   Warranty conditions, liability, AND support -
      IF the application has been made available free OF charge, the following applies:
      * We DO NOT provide a warranty FOR Any OF the information contained in this document.
      * All other rights AND claims against Siemens AG irrespective OF legal basis are excluded. In particular claims FOR damages against Siemens AG 
      in the CASE OF Product outage, downtime, loss OF profit, either directly, indirectly OR consequential damage are excluded.
      * This does NOT apply when liability is compulsory BY law, e. g. in the CASE OF the Product liability act, premeditation, an act OF gross negligence 
      BY superiors AND managerial staff OF Siemens AG OR in cases OF fraudulent concealment OF defects.
      * This limitation OF liability also applies TO sub-contractors, suppliers, delegates, superiors AND managerial staff OF Siemens AG.
      German law shall apply TO this agreement FOR customers with head offices in Germany; Swiss law FOR customers with head offices outside Germany. 
      Application OF the United Nations Convention on Contracts FOR the International Sale OF Goods as OF 11.04.1980 (CISG) is excluded.
   *)

   // ===========================================================================
   //  Begin the LOGIC section:
   //  

    #temp_UDint := 0;

   IF IS_ARRAY(#Array_ToBe_Sized) THEN                             // Is this a valid array?
       #temp_UDint := CountOfElements(#Array_ToBe_Sized);          // Determine the length of the array...
   END_IF;

   #ArraySize := UDINT_TO_INT(#temp_UDint);

   // End of Main Logic Section 
   ENO := true;   // Set the ENO output
END_FUNCTION

(* ===== HMI "HMI_RT_1" =====
system functions are stored by id; their names below are inferred from use

HMI tags "Default tag table"
   "bo_PreviousPage_pressed" : Bool, internal
   "bo_NextPage_pressed" : Bool, internal

ScreenModuleEditorView "typ_ThirdLevelNavigation" 165x50
   Button "Btn_NextPage" at 115,0 size 50x50; TextOff 'Text'; PictureOff "Right_transparent_48x48"
      on Press: function_b14e0dd5("bo_NextPage_pressed", 0)
      Appearance <- "bo_NextPage_pressed"
   Button "btn_PreviousPage" at 0,0 size 50x50; TextOff 'Text'; PictureOff "Left_transparent_48x48"
      on Press: function_b14e0dd5("bo_PreviousPage_pressed", 0)
      Appearance <- "bo_PreviousPage_pressed"
   TextField "txt_actualID" at 55,11 size 28x27; Text '11'
   TextField "txt_maximum _ID" at 82,11 size 28x27; Text '11'
   TextField "txt_Backslash" at 76,11 size 14x27; Text '/'
   GraphicView "pic_transparent_previous" at 0,0 size 50x50; Picture "btn-disabled-50x50"
      Visibility <- "bo_PreviousActive"
   GraphicView "pic_transparent_next" at 115,0 size 50x50; Picture "btn-disabled-50x50"
      Visibility <- "bo_NextActive"
*)

(* ===== HMI "HMI_RT_1" =====

ScreenModuleEditorView "fcpOmacTime" 490x26
   IOField "valOutputModeName" at 0,0 size 151x26; FormatPattern ??????????????????
      ProcessValue <- "ModeName"
   IOField "valOutputCurrentTime" at 150,0 size 101x26; FormatPattern 999999999
      ProcessValue <- "CurrentTime"
   IOField "ValOutputCumulativeTime" at 250,0 size 101x26; FormatPattern 999999999
      ProcessValue <- "CumulativeTime"
   Bar "valOutputCumuliativeTimePercent" at 355,5 size 131x16; MinimumValue 0; MaximumValue 100
      ProcessValue <- "CumulativeTime"
      MaximumValue <- "TimeOverAll"
*)

(* ===== HMI "HMI_RT_1" =====
system functions are stored by id; their names below are inferred from use

HMI tags "Standard-Variablentabelle"
   "bo_Topic01BtnPressed" : Bool, internal
   "bo_Topic02BtnPressed" : Bool, internal
   "bo_Topic03BtnPressed" : Bool, internal
   "bo_Topic04BtnPressed" : Bool, internal
   "bo_Topic05BtnPressed" : Bool, internal
   "bo_Topic06BtnPressed" : Bool, internal
   "bo_Topic07BtnPressed" : Bool, internal
   "bo_Topic08BtnPressed" : Bool, internal
   "bo_Topic09BtnPressed" : Bool, internal
   "bo_Topic10BtnPressed" : Bool, internal
   "bo_Topic11BtnPressed" : Bool, internal
   "bo_Topic12BtnPressed" : Bool, internal
   "bo_Topic13BtnPressed" : Bool, internal
   "bo_Topic14BtnPressed" : Bool, internal
   "bo_Topic15BtnPressed" : Bool, internal
   "bo_Topic16BtnPressed" : Bool, internal
   "bo_Topic17BtnPressed" : Bool, internal
   "bo_Topic18BtnPressed" : Bool, internal
   "bo_Topic19BtnPressed" : Bool, internal
   "bo_Topic20BtnPressed" : Bool, internal
   "bo_Topic21BtnPressed" : Bool, internal
   "bo_Topic22BtnPressed" : Bool, internal
   "bo_Topic23BtnPressed" : Bool, internal
   "bo_Topic24BtnPressed" : Bool, internal
   "i16_configReg" : Int, internal   // Combination of actual showed LvL and input configuration of used Register; To show active Register
   "i16_LvL_Shown" : Int, internal   // number of actual showed LvL
   "i16_SaveScreenNo" : Int, internal   // Save actual Screen Number
   "i16_RegShown" : Int, internal   // Combination of actual active Register and actual active LvL; to show the active Register
   "bo_NextTopicLvL1" : Int, internal
   "i16_InputScreenID" : Int, internal   // help Variable
   "i16_Input_maxReg" : Int, internal   // help Variable
   "i16_RegNo" : Int, internal   // Active Register number;Value 1-24
   "bo_PreviousPageBtnPressed" : Bool, internal

ScreenModuleEditorView "fcpSecondLevelNavigation" 1270x615
   Rectangle "rec_Topic_001.0" at 207,42 size 1063x62
      Visibility <- "i16_RegShown"
   Rectangle "rec_Topic_002.0" at 207,109 size 1063x62
      Visibility <- "i16_RegShown"
   Rectangle "rec_Topic_003.0" at 207,176 size 1063x62
      Visibility <- "i16_RegShown"
   Rectangle "rec_Topic_004.0" at 207,243 size 1063x62
      Visibility <- "i16_RegShown"
   Rectangle "rec_Topic_005.0" at 207,310 size 1063x62
      Visibility <- "i16_RegShown"
   Rectangle "rec_Topic_006.0" at 207,377 size 1063x62
      Visibility <- "i16_RegShown"
   Rectangle "rec_Topic_007.0" at 207,444 size 1063x62
      Visibility <- "i16_RegShown"
   Rectangle "rec_Topic_008.0" at 207,511 size 1063x62
      Visibility <- "i16_RegShown"
   TextField "txt_Topic_001.0_Textfield" at 1100,42 size 170x62; Text 'Thema 001.0 / Topic 001.0'
      Visibility <- "i16_configReg"
      Appearance <- "i16_RegShown"
   Button "btn_Topic_001.0_Button" at 1100,42 size 170x62; TextOff 'Text'
      on Release: "sub_TabLvL"()
      on Press: function_b14e0dd5("bo_Topic01BtnPressed", 0)
      Visibility <- "i16_configReg"
   TextField "txt_Topic_002.0_Textfield" at 1100,109 size 170x62; Text 'Thema 002.0 / Topic 002.0'
      Visibility <- "i16_configReg"
      Appearance <- "i16_RegShown"
   Button "btn_Topic_002.0_Button" at 1100,109 size 170x62; TextOff 'Text'
      on Release: "sub_TabLvL"()
      on Press: function_b14e0dd5("bo_Topic02BtnPressed", 0)
      Visibility <- "i16_configReg"
   TextField "txt_Topic_003.0_Textfield" at 1100,176 size 170x62; Text 'Thema 003.0 / Topic 003.0'
      Visibility <- "i16_configReg"
      Appearance <- "i16_RegShown"
   Button "btn_Topic_003.0_Button" at 1100,176 size 170x62; TextOff 'Text'
      on Release: "sub_TabLvL"()
      on Press: function_b14e0dd5("bo_Topic03BtnPressed", 0)
      Visibility <- "i16_configReg"
   TextField "txt_Topic_004.0_Textfield" at 1100,243 size 170x62; Text 'Thema 004.0 / Topic 004.0'
      Visibility <- "i16_configReg"
      Appearance <- "i16_RegShown"
   Button "btn_Topic_004.0_Button" at 1100,243 size 170x62; TextOff 'Text'
      on Release: "sub_TabLvL"()
      on Press: function_b14e0dd5("bo_Topic04BtnPressed", 0)
      Visibility <- "i16_configReg"
   TextField "txt_Topic_005.0_Textfield" at 1100,310 size 170x62; Text 'Thema 005.0 / Topic 005.0'
      Visibility <- "i16_configReg"
      Appearance <- "i16_RegShown"
   Button "btn_Topic_005.0_Button" at 1100,310 size 170x62; TextOff 'Text'
      on Release: "sub_TabLvL"()
      on Press: function_b14e0dd5("bo_Topic05BtnPressed", 0)
      Visibility <- "i16_configReg"
   TextField "txt_Topic_006.0_Textfield" at 1100,377 size 170x62; Text 'Thema 006.0 / Topic 006.0 / Topic 005.0'
      Visibility <- "i16_configReg"
      Appearance <- "i16_RegShown"
   Button "btn_Topic_006.0_Button" at 1100,377 size 170x62; TextOff 'Text'
      on Release: "sub_TabLvL"()
      on Press: function_b14e0dd5("bo_Topic06BtnPressed", 0)
      Visibility <- "i16_configReg"
   TextField "txt_Topic_007.0_Textfield" at 1100,444 size 170x62; Text 'Thema 007.0 / Topic 007.0 / Topic 005.0'
      Visibility <- "i16_configReg"
      Appearance <- "i16_RegShown"
   Button "btn_Topic_007.0_Button" at 1100,444 size 170x62; TextOff 'Text'
      on Release: "sub_TabLvL"()
      on Press: function_b14e0dd5("bo_Topic07BtnPressed", 0)
      Visibility <- "i16_configReg"
   TextField "txt_Topic_008.0_Textfield" at 1100,511 size 170x62; Text 'Thema 007.0 / Topic 008.0 / Topic 005.0'
      Visibility <- "i16_configReg"
      Appearance <- "i16_RegShown"
   Button "btn_Topic_008.0_Button" at 1100,511 size 170x62; TextOff 'Text'
      on Release: "sub_TabLvL"()
      on Press: function_b14e0dd5("bo_Topic08BtnPressed", 0)
      Visibility <- "i16_configReg"
   Rectangle "rec_Topic_001.0_RectangleLight" at 1100,42 size 170x62
      Visibility <- "i16_configReg"
      Appearance <- "bo_Topic01BtnPressed"
   Rectangle "rec_Topic_002.0_RectangleLight" at 1100,109 size 170x62
      Visibility <- "i16_configReg"
      Appearance <- "bo_Topic02BtnPressed"
   Rectangle "rec_Topic_003.0_RectangleLight" at 1100,176 size 170x62
      Visibility <- "i16_configReg"
      Appearance <- "bo_Topic03BtnPressed"
   Rectangle "rec_Topic_004.0_RectangleLight" at 1100,243 size 170x62
      Visibility <- "i16_configReg"
      Appearance <- "bo_Topic04BtnPressed"
   Rectangle "rec_Topic_005.0_RectangleLight" at 1100,310 size 170x62
      Visibility <- "i16_configReg"
      Appearance <- "bo_Topic05BtnPressed"
   Rectangle "rec_Topic_006.0_RectangleLight" at 1100,377 size 170x62
      Visibility <- "i16_configReg"
      Appearance <- "bo_Topic06BtnPressed"
   Rectangle "rec_Topic_007.0_RectangleLight" at 1100,444 size 170x62
      Visibility <- "i16_configReg"
      Appearance <- "bo_Topic07BtnPressed"
   Rectangle "rec_Topic_008.0_RectangleLight" at 1100,511 size 170x62
      Visibility <- "i16_configReg"
      Appearance <- "bo_Topic08BtnPressed"
   Rectangle "rec_Topic_009.0_RectangleLight" at 1100,42 size 170x62
      Visibility <- "i16_configReg"
      Appearance <- "bo_Topic09BtnPressed"
   Rectangle "rec_Topic_010.0_RectangleLight" at 1100,109 size 170x62
      Visibility <- "i16_configReg"
      Appearance <- "bo_Topic10BtnPressed"
   Rectangle "rec_Topic_011.0_RectangleLight" at 1100,176 size 170x62
      Visibility <- "i16_configReg"
      Appearance <- "bo_Topic11BtnPressed"
   Rectangle "rec_Topic_012.0_RectangleLight" at 1100,243 size 170x62
      Visibility <- "i16_configReg"
      Appearance <- "bo_Topic12BtnPressed"
   Rectangle "rec_Topic_013.0_RectangleLight" at 1100,310 size 170x62
      Visibility <- "i16_configReg"
      Appearance <- "bo_Topic13BtnPressed"
   Rectangle "rec_Topic_014.0_RectangleLight" at 1100,377 size 170x62
      Visibility <- "i16_configReg"
      Appearance <- "bo_Topic14BtnPressed"
   Rectangle "rec_Topic_015.0_RectangleLight" at 1100,444 size 170x62
      Visibility <- "i16_configReg"
      Appearance <- "bo_Topic15BtnPressed"
   Rectangle "rec_Topic_016.0_RectangleLight" at 1100,511 size 170x62
      Visibility <- "i16_configReg"
      Appearance <- "bo_Topic16BtnPressed"
   Rectangle "rec_Topic_009.0" at 207,42 size 1063x62
      Visibility <- "i16_RegShown"
   Rectangle "rec_Topic_010.0" at 207,109 size 1063x62
      Visibility <- "i16_RegShown"
   Rectangle "rec_Topic_011.0" at 207,176 size 1063x62
      Visibility <- "i16_RegShown"
   Rectangle "rec_Topic_012.0" at 207,243 size 1063x62
      Visibility <- "i16_RegShown"
   Rectangle "rec_Topic_013.0" at 207,310 size 1063x62
      Visibility <- "i16_RegShown"
   Rectangle "rec_Topic_014.0" at 207,377 size 1063x62
      Visibility <- "i16_RegShown"
   Rectangle "rec_Topic_015.0" at 207,444 size 1063x62
      Visibility <- "i16_RegShown"
   Rectangle "rec_Topic_016.0" at 207,511 size 1063x62
      Visibility <- "i16_RegShown"
   Rectangle "rec_Topic_017.0_RectangleLight" at 1100,42 size 170x62
      Visibility <- "i16_configReg"
      Appearance <- "bo_Topic17BtnPressed"
   Rectangle "rec_Topic_018.0_RectangleLight" at 1100,109 size 170x62
      Visibility <- "i16_configReg"
      Appearance <- "bo_Topic18BtnPressed"
   Rectangle "rec_Topic_019.0_RectangleLight" at 1100,176 size 170x62
      Visibility <- "i16_configReg"
      Appearance <- "bo_Topic19BtnPressed"
   Rectangle "rec_Topic_020.0_RectangleLight" at 1100,243 size 170x62
      Visibility <- "i16_configReg"
      Appearance <- "bo_Topic20BtnPressed"
   Rectangle "rec_Topic_021.0_RectangleLight" at 1100,310 size 170x62
      Visibility <- "i16_configReg"
      Appearance <- "bo_Topic21BtnPressed"
   Rectangle "rec_Topic_022.0_RectangleLight" at 1100,377 size 170x62
      Visibility <- "i16_configReg"
      Appearance <- "bo_Topic22BtnPressed"
   Rectangle "rec_Topic_023.0_RectangleLight" at 1100,444 size 170x62
      Visibility <- "i16_configReg"
      Appearance <- "bo_Topic23BtnPressed"
   Rectangle "rec_Topic_024.0_RectangleLight" at 1100,511 size 170x62
      Visibility <- "i16_configReg"
      Appearance <- "bo_Topic24BtnPressed"
   Rectangle "rec_Topic_017.0" at 207,42 size 1063x62
      Visibility <- "i16_RegShown"
   Rectangle "rec_Topic_018.0" at 207,109 size 1063x62
      Visibility <- "i16_RegShown"
   Rectangle "rec_Topic_019.0" at 207,176 size 1063x62
      Visibility <- "i16_RegShown"
   Rectangle "rec_Topic_020.0" at 207,243 size 1063x62
      Visibility <- "i16_RegShown"
   Rectangle "rec_Topic_021.0" at 207,310 size 1063x62
      Visibility <- "i16_RegShown"
   Rectangle "rec_Topic_022.0" at 207,377 size 1063x62
      Visibility <- "i16_RegShown"
   Rectangle "rec_Topic_023.0" at 207,444 size 1063x62
      Visibility <- "i16_RegShown"
   Rectangle "rec_Topic_024.0" at 207,511 size 1063x62
      Visibility <- "i16_RegShown"
   TextField "txt_Topic_009.0_Textfield" at 1100,42 size 170x62; Text 'Thema 001.0 / Topic 009.0 / Topic 001.0'
      Visibility <- "i16_configReg"
      Appearance <- "i16_RegShown"
   Button "btn_Topic_009.0_Button" at 1100,42 size 170x62; TextOff 'Text'
      on Release: "sub_TabLvL"()
      on Press: function_b14e0dd5("bo_Topic09BtnPressed", 0)
      Visibility <- "i16_configReg"
   TextField "txt_Topic_010.0_Textfield" at 1100,109 size 170x62; Text 'Thema 002.0 / Topic 010.0 / Topic 002.0'
      Visibility <- "i16_configReg"
      Appearance <- "i16_RegShown"
   Button "btn_Topic_010.0_Button" at 1100,109 size 170x62; TextOff 'Text'
      on Release: "sub_TabLvL"()
      on Press: function_b14e0dd5("bo_Topic10BtnPressed", 0)
      Visibility <- "i16_configReg"
   TextField "txt_Topic_011.0_Textfield" at 1100,176 size 170x62; Text 'Thema 003.0 / Topic 011.0 / Topic 003.0'
      Visibility <- "i16_configReg"
      Appearance <- "i16_RegShown"
   Button "btn_Topic_011.0_Button" at 1100,176 size 170x62; TextOff 'Text'
      on Release: "sub_TabLvL"()
      on Press: function_b14e0dd5("bo_Topic11BtnPressed", 0)
      Visibility <- "i16_configReg"
   TextField "txt_Topic_012.0_Textfield" at 1100,243 size 170x62; Text 'Thema 004.0 / Topic 012.0 / Topic 004.0'
      Visibility <- "i16_configReg"
      Appearance <- "i16_RegShown"
   Button "btn_Topic_012.0_Button" at 1100,243 size 170x62; TextOff 'Text'
      on Release: "sub_TabLvL"()
      on Press: function_b14e0dd5("bo_Topic12BtnPressed", 0)
      Visibility <- "i16_configReg"
   TextField "txt_Topic_013.0_Textfield" at 1100,310 size 170x62; Text 'Thema 005.0 / Topic 013.0 / Topic 005.0'
      Visibility <- "i16_configReg"
      Appearance <- "i16_RegShown"
   Button "btn_Topic_013.0_Button" at 1100,310 size 170x62; TextOff 'Text'
      on Release: "sub_TabLvL"()
      on Press: function_b14e0dd5("bo_Topic13BtnPressed", 0)
      Visibility <- "i16_configReg"
   TextField "txt_Topic_014.0_Textfield" at 1100,377 size 170x62; Text 'Thema 006.0 / Topic 014.0 / Topic 005.0'
      Visibility <- "i16_configReg"
      Appearance <- "i16_RegShown"
   Button "btn_Topic_014.0_Button" at 1100,377 size 170x62; TextOff 'Text'
      on Release: "sub_TabLvL"()
      on Press: function_b14e0dd5("bo_Topic14BtnPressed", 0)
      Visibility <- "i16_configReg"
   TextField "txt_Topic_015.0_Textfield" at 1100,444 size 170x62; Text 'Thema 007.0 / Topic 015.0 / Topic 005.0'
      Visibility <- "i16_configReg"
      Appearance <- "i16_RegShown"
   Button "btn_Topic_015.0_Button" at 1100,444 size 170x62; TextOff 'Text'
      on Release: "sub_TabLvL"()
      on Press: function_b14e0dd5("bo_Topic15BtnPressed", 0)
      Visibility <- "i16_configReg"
   TextField "txt_Topic_016.0_Textfield" at 1100,511 size 170x62; Text 'Thema 007.0 / Topic 016.0 / Topic 005.0'
      Visibility <- "i16_configReg"
      Appearance <- "i16_RegShown"
   Button "btn_Topic_016.0_Button" at 1100,511 size 170x62; TextOff 'Text'
      on Release: "sub_TabLvL"()
      on Press: function_b14e0dd5("bo_Topic16BtnPressed", 0)
      Visibility <- "i16_configReg"
   TextField "txt_Topic_017.0_Textfield" at 1100,42 size 170x62; Text 'Thema 001.0 / Topic 017.0 / Topic 001.0'
      Visibility <- "i16_configReg"
      Appearance <- "i16_RegShown"
   Button "btn_Topic_017.0_Button" at 1100,42 size 170x62; TextOff 'Text'
      on Release: "sub_TabLvL"()
      on Press: function_b14e0dd5("bo_Topic17BtnPressed", 0)
      Visibility <- "i16_configReg"
   TextField "txt_Topic_018.0_Textfield" at 1100,109 size 170x62; Text 'Thema 002.0 / Topic 018.0 / Topic 002.0'
      Visibility <- "i16_configReg"
      Appearance <- "i16_RegShown"
   Button "btn_Topic_018.0_Button" at 1100,109 size 170x62; TextOff 'Text'
      on Release: "sub_TabLvL"()
      on Press: function_b14e0dd5("bo_Topic18BtnPressed", 0)
      Visibility <- "i16_configReg"
   TextField "txt_Topic_019.0_Textfield" at 1100,176 size 170x62; Text 'Thema 003.0 / Topic 019.0 / Topic 003.0'
      Visibility <- "i16_configReg"
      Appearance <- "i16_RegShown"
   Button "btn_Topic_019.0_Button" at 1100,176 size 170x62; TextOff 'Text'
      on Release: "sub_TabLvL"()
      on Press: function_b14e0dd5("bo_Topic19BtnPressed", 0)
      Visibility <- "i16_configReg"
   TextField "txt_Topic_020.0_Textfield" at 1100,243 size 170x62; Text 'Thema 004.0 / Topic 020.0 / Topic 004.0'
      Visibility <- "i16_configReg"
      Appearance <- "i16_RegShown"
   Button "btn_Topic_020.0_Button" at 1100,243 size 170x62; TextOff 'Text'
      on Release: "sub_TabLvL"()
      on Press: function_b14e0dd5("bo_Topic20BtnPressed", 0)
      Visibility <- "i16_configReg"
   TextField "txt_Topic_021.0_Textfield" at 1100,310 size 170x62; Text 'Thema 005.0 / Topic 021.0 / Topic 005.0'
      Visibility <- "i16_configReg"
      Appearance <- "i16_RegShown"
   Button "btn_Topic_021.0_Button" at 1100,310 size 170x62; TextOff 'Text'
      on Release: "sub_TabLvL"()
      on Press: function_b14e0dd5("bo_Topic21BtnPressed", 0)
      Visibility <- "i16_configReg"
   TextField "txt_Topic_022.0_Textfield" at 1100,377 size 170x62; Text 'Thema 006.0 / Topic 022.0 / Topic 005.0'
      Visibility <- "i16_configReg"
      Appearance <- "i16_RegShown"
   Button "btn_Topic_022.0_Button" at 1100,377 size 170x62; TextOff 'Text'
      on Release: "sub_TabLvL"()
      on Press: function_b14e0dd5("bo_Topic22BtnPressed", 0)
      Visibility <- "i16_configReg"
   TextField "txt_Topic_023.0_Textfield" at 1100,444 size 170x62; Text 'Thema 007.0 / Topic 023.0 / Topic 005.0'
      Visibility <- "i16_configReg"
      Appearance <- "i16_RegShown"
   Button "btn_Topic_023.0_Button" at 1100,444 size 170x62; TextOff 'Text'
      on Release: "sub_TabLvL"()
      on Press: function_b14e0dd5("bo_Topic23BtnPressed", 0)
      Visibility <- "i16_configReg"
   TextField "txt_Topic_024.0_Textfield" at 1100,511 size 170x62; Text 'Thema 007.0 / Topic 024.0 / Topic 005.0'
      Visibility <- "i16_configReg"
      Appearance <- "i16_RegShown"
   Button "btn_Topic_024.0_Button" at 1100,511 size 170x62; TextOff 'Text'
      on Release: "sub_TabLvL"()
      on Press: function_b14e0dd5("bo_Topic24BtnPressed", 0)
      Visibility <- "i16_configReg"
   Rectangle "rec_Topic_008.0_RectangleLight_1" at 1100,578 size 170x37
      Appearance <- "bo_NextTopicLvL1"
   GraphicView "pic_ArrowDown" at 1161,578 size 48x37; Picture "Down_transparent_48x48"
   Button "btn_Topic_008.0_Button_1" at 1100,578 size 170x37; TextOff 'Text'
      on Release: function_dd21b452("i16_LvL_Shown", 1); SetTag("i16_Input_maxReg", "i16_MaxTopics"); "sub_TabLvL"()
      on Press: function_b14e0dd5("bo_NextTopicLvL1", 0)
      ObjectEnable <- "i16_LvL_Shown"
   Rectangle "rec_Topic_008.0_RectangleLight_2" at 1100,0 size 170x37
      Visibility <- "i16_MaxTopics"
      Appearance <- "bo_PreviousPageBtnPressed"
   GraphicView "pic_ArrowUp" at 1161,0 size 48x37; Picture "Line-Up_transparent_48x48"
      Visibility <- "i16_MaxTopics"
   Button "btn_Topic_008.0_Button_2" at 1100,0 size 170x37; TextOff 'Text'
      on Release: function_b9b71300("i16_LvL_Shown", 1); "sub_TabLvL"()
      on Press: function_b14e0dd5("bo_PreviousPageBtnPressed", 0)
      Visibility <- "i16_MaxTopics"
      ObjectEnable <- "i16_LvL_Shown"
   Rectangle "rec_Topic_008.0_RectangleLight_4" at 1100,578 size 170x37
      Visibility <- "i16_LvL_Shown"
      Appearance <- "bo_NextTopicLvL1"
   GraphicView "pic_ArrowDown_1" at 1161,578 size 48x37; Picture "Down_transparent_48x48"
      Visibility <- "i16_LvL_Shown"
   Button "btn_Topic_008.0_Button_3" at 1100,578 size 170x37; TextOff 'Text'
      on Release: function_dd21b452("i16_LvL_Shown", 1); "sub_TabLvL"()
      on Press: function_b14e0dd5("bo_NextTopicLvL1", 0)
      Visibility <- "i16_LvL_Shown"
      ObjectEnable <- "i16_LvL_Shown"
   GraphicView "pic_Transparent_PreviousScreen" at 1100,0 size 170x37; Picture "btn-disabled-170x31"
      Visibility <- "i16_LvL_Shown"
   GraphicView "pic_Transparent_NextPageLvL1" at 1100,578 size 170x37; Picture "btn-disabled-170x31"
      Visibility <- "i16_configReg"
   GraphicView "pic_Transparent_NextPageLvL2" at 1100,578 size 170x37; Picture "btn-disabled-170x31"
      Visibility <- "i16_configReg"
   GraphicView "pic_Transparent_NextPageLvL3" at 1100,578 size 170x37; Picture "btn-disabled-170x31"
      Visibility <- "i16_configReg"

VB script "sub_TabLvL"
   'Declaration
   Dim NoMainTopic, ScreenID, actRegNo
   
   
   ScreenID = SmartTags("i16_CurScreenID")
   'Check if 1.Time Script
   If SmartTags("i16_LvL_Shown")= 0 Then
   	SmartTags("i16_LvL_Shown")=1
   End If 
   'check if new Screen
   If SmartTags("i16_SaveScreenNo")=SmartTags("i16_CurScreenID") Then 'SmartTags("i16_InputScreenID")Then 
   	'No new Screen
   Else
   	'New Screen open
   	 	
   	'check active Register	 
   		NoMainTopic = 0
   		'Screen ID to internal Variable
   		ScreenID =SmartTags("i16_CurScreenID") 'SmartTags("i16_InputScreenID")
   		'Save ScreenID
   		SmartTags("i16_SaveScreenNo")=SmartTags("i16_CurScreenID") 'SmartTags("i16_InputScreenID")
   		'Seperate ScreenID: Filter MainTopic
   		While ScreenID > 1000
   			NoMainTopic = NoMainTopic + 1 ' Main Topic - Machine COntrol etc.
   			ScreenID = ScreenID -1000
   		Wend 
   	
   		'initialise actual Register number
   		actRegNo = 0 
   		
   		'Seperate Screen ID: Which Register is active ; possible Value 1-24
   		While ScreenID >= 0 
   			ScreenID =  ScreenID - 40
   			actRegNo = actRegNo + 1
   		Wend
   		
   		'Save active Register Number
   		SmartTags("i16_RegNo")= 	actRegNo
   	'Set actual Secundary Level number 
   	If actRegNo < 9 Then ' 1-8=LvL1
   		SmartTags("i16_LvL_Shown")= 1
   	End If 
   	
   	If actRegNo > 8 And actRegNo<17 Then '9-16=LvL2
   		SmartTags("i16_LvL_Shown")= 2
   	End If 
   	
   	If actRegNo > 16 Then ' 17-24=LvL3
   		SmartTags("i16_LvL_Shown")= 3
   	End If 
   End If 
   			
   'code the Variable 'i16_RegShown' with the actual shown LvL and the actual shown Register
   SmartTags("i16_RegShown")= SmartTags("i16_LvL_Shown")* 100 + SmartTags("i16_RegNo")
   
   '----------------------------------------------------
   
   'check configuration of used Register
   SmartTags("i16_configReg") =SmartTags("i16_LvL_Shown") * 100 + SmartTags("i16_MaxTopics") 'SmartTags("i16_Input_maxReg")
   ' 1. no := LvL; 2.& 3. := configuration of Tabs 
   
   'LvL+100 + sekundary Lvl aktive
   
   
   '	
*)

(* ===== HMI "HMI_RT_1" =====
system functions are stored by id; their names below are inferred from use

HMI tags "Standard-Variablentabelle"
   "bo_MachineControlBtnPressed" : Bool, internal
   "bo_SettingsBtnPressed" : Bool, internal
   "bo_Alarm&EventsBtnPressed" : Bool, internal
   "bo_StatisticsBtnPressed" : Bool, internal
   "bo_ManualBtnPressed" : Bool, internal
   "bo_DiagnosticsBtnPressed" : Bool, internal
   "bo_FormatBtnPressed" : Bool, internal
   "bo_LogonBtnPressed" : Bool, internal
   "bo_PreviousScreenBtnPressed" : Bool, internal

ScreenModuleEditorView "fcpBottomBar" 1270x85
   Rectangle "rec_MachineControlSelected" at 0,0 size 152x11
      Visibility <- "ScreenNo"
   Rectangle "rec_SettingsSelected" at 157,0 size 152x11
      Visibility <- "ScreenNo"
   Rectangle "rec_Alarm&EventsSelected" at 314,0 size 152x11
      Visibility <- "ScreenNo"
   Rectangle "rec_DiagnosticsSelected" at 471,0 size 152x11
      Visibility <- "ScreenNo"
   Rectangle "rec_FormatsSelected" at 628,0 size 153x11
      Visibility <- "ScreenNo"
   Rectangle "rec_MachineControl" at 0,12 size 152x73
      Appearance <- "bo_MachineControlBtnPressed"
   Rectangle "rec_Settings" at 157,12 size 152x73
      Appearance <- "bo_SettingsBtnPressed"
   Rectangle "rec_Alarm&Events" at 314,12 size 152x73
      Appearance <- "bo_Alarm&EventsBtnPressed"
   Rectangle "rec_Diagnostics" at 471,12 size 152x73
      Appearance <- "bo_DiagnosticsBtnPressed"
   Rectangle "rec_Formats" at 628,12 size 153x73
      Appearance <- "bo_FormatBtnPressed"
   Rectangle "rec_PreviousScreen" at 1100,12 size 83x73
      Appearance <- "bo_PreviousScreenBtnPressed"
   Rectangle "rec_Logon" at 1188,12 size 82x73
      Appearance <- "bo_LogonBtnPressed"
   TextField "txt_MachineControl" at 0,12 size 152x73; Text 'Maschine / Machine control / Topic 001.1'
   TextField "txt_Settings" at 157,12 size 152x73; Text 'Einstellungen / Settings / Topic 001.1'
   TextField "txt_Alarm&Events" at 314,12 size 152x73; Text 'Meldungen / Alarm & Events / Topic 001.1'
   TextField "txt_Diagnostics" at 471,12 size 152x73; Text 'Diagnose / Diagnostics / Topic 001.1'
   TextField "txt_Formats" at 628,12 size 153x73; Text 'Formate / Formats / Topic 001.1'
   TextField "txt_PrevousScreen" at 1100,12 size 83x73; Text 'Zurück / Back / Topic 001.1'
   TextField "txt_Logon" at 1188,12 size 82x73; Text 'Logon / Topic 001.1'
   GraphicView "pic_MachineControl" at 53,36 size 48x48; Picture "Production_transparent_48x48"
   GraphicView "pic_Settings" at 210,36 size 48x48; Picture "Setup_transparent_48x48"
   GraphicView "pic_Alarm&Events" at 367,36 size 48x48; Picture "Alarm_transparent_48x48"
   GraphicView "pic_Diagnostics" at 524,36 size 48x48; Picture "Diagnostics_transparent_48x48"
   GraphicView "pic_Formats" at 681,36 size 48x48; Picture "InsertLine_transparent_48x48"
   GraphicView "pic_PreviousScreen" at 1118,36 size 48x48; Picture "Back_transparent_48x48[1]"
   GraphicView "pic_Login" at 1206,36 size 48x48; Picture "Login_transparent_48x48[1]"
   Button "btn_MachineControl" at 0,12 size 152x73; TextOff 'Text'
      on Press: function_b14e0dd5("bo_MachineControlBtnPressed", 0)
   Button "btn_Settings" at 157,12 size 152x73; TextOff 'Text'
      on Press: function_b14e0dd5("bo_SettingsBtnPressed", 0)
   Button "btn_Alarm&Events" at 314,12 size 152x73; TextOff 'Text'
      on Press: function_b14e0dd5("bo_Alarm&EventsBtnPressed", 0)
   Button "btn_Diagnostics" at 471,12 size 152x73; TextOff 'Text'
      on Press: function_b14e0dd5("bo_DiagnosticsBtnPressed", 0)
   Button "btn_Formats" at 628,12 size 153x73; TextOff 'Text'
      on Press: function_b14e0dd5("bo_FormatBtnPressed", 0)
   Button "btn_PreviousScreen" at 1100,12 size 83x73; TextOff 'Text'
      on Press: function_b14e0dd5("bo_PreviousScreenBtnPressed", 0)
   Button "btn_Logon" at 1188,12 size 82x73; TextOff 'Text'
      on Press: function_b14e0dd5("bo_LogonBtnPressed", 0)
*)

(* ===== HMI "HMI_RT_1" =====

ScreenModuleEditorView "fcpEvent_Status_AlarmsWarning_withValue" 1030x51
   IOField "valOutputTop_ID" at 0,0 size 56x26; FormatPattern 99999
      ProcessValue <- "1_Top_PropertiesTag.ID"
      Appearance <- "1_Top_PropertiesTag.ID"
   IOField "valOutputTop_Value" at 55,0 size 56x26; FormatPattern 99999
      ProcessValue <- "1_Top_PropertiesTag.Value"
      Appearance <- "1_Top_PropertiesTag.ID"
   IOField "valOutputTop_Category" at 110,0 size 31x26; FormatPattern 99
      ProcessValue <- "1_Top_PropertiesTag.Category"
      Appearance <- "1_Top_PropertiesTag.ID"
   IOField "valOutputTop_Message" at 140,0 size 491x26; FormatPattern ??????????????????????????????????????????????????
      ProcessValue <- "1_Top_PropertiesTag.Message"
      Appearance <- "1_Top_PropertiesTag.ID"
   IOField "valOutputTop_DateTime" at 630,0 size 201x26
      Appearance <- "1_Top_PropertiesTag.ID"
      ProcessValue <- "1_Top_PropertiesTag.DateTimeDTL"
   IOField "valOutputTop_AckDateTime" at 830,0 size 200x26
      Appearance <- "1_Top_PropertiesTag.ID"
      ProcessValue <- "1_Top_PropertiesTag.AckDateTimeDTL"
   IOField "valOutputBottom_ID" at 0,25 size 56x26; FormatPattern 99999
      ProcessValue <- "2_Bottom_PropertiesTag.ID"
      Appearance <- "2_Bottom_PropertiesTag.ID"
   IOField "valOutputBottom_Value" at 55,25 size 56x26; FormatPattern 99999
      ProcessValue <- "2_Bottom_PropertiesTag.Value"
      Appearance <- "2_Bottom_PropertiesTag.ID"
   IOField "valOutputBottom_Category" at 110,25 size 31x26; FormatPattern 99
      ProcessValue <- "2_Bottom_PropertiesTag.Category"
      Appearance <- "2_Bottom_PropertiesTag.ID"
   IOField "valOutputBottom_Message" at 140,25 size 491x26; FormatPattern ??????????????????????????????????????????????????
      ProcessValue <- "2_Bottom_PropertiesTag.Message"
      Appearance <- "2_Bottom_PropertiesTag.ID"
   IOField "valOutputBottom_DateTime" at 630,25 size 201x26
      Appearance <- "2_Bottom_PropertiesTag.ID"
      ProcessValue <- "2_Bottom_PropertiesTag.DateTimeDTL"
   IOField "valOutputBottom_AckDateTime" at 830,25 size 200x26
      Appearance <- "2_Bottom_PropertiesTag.ID"
      ProcessValue <- "2_Bottom_PropertiesTag.AckDateTimeDTL"
*)

(* ===== HMI "HMI_RT_1" =====

ScreenModuleEditorView "fcpEvent_Status_AlarmsWarning" 1030x51
   IOField "valOutputTop_ID" at 0,0 size 56x26; FormatPattern 99999
      ProcessValue <- "1_Top_PropertiesTag.ID"
      Appearance <- "1_Top_PropertiesTag.ID"
   IOField "valOutputTop_Category" at 55,0 size 31x26; FormatPattern 99
      ProcessValue <- "1_Top_PropertiesTag.Category"
      Appearance <- "1_Top_PropertiesTag.ID"
   IOField "valOutputTop_Message" at 85,0 size 546x26; FormatPattern ??????????????????????????????????????????????????
      ProcessValue <- "1_Top_PropertiesTag.Message"
      Appearance <- "1_Top_PropertiesTag.ID"
   IOField "valOutputTop_DateTime" at 630,0 size 201x26
      Appearance <- "1_Top_PropertiesTag.ID"
      ProcessValue <- "1_Top_PropertiesTag.DateTimeDTL"
   IOField "valOutputTop_AckDateTime" at 830,0 size 200x26
      Appearance <- "1_Top_PropertiesTag.ID"
      ProcessValue <- "1_Top_PropertiesTag.AckDateTimeDTL"
   IOField "valOutputBottom_ID" at 0,25 size 56x26; FormatPattern 99999
      ProcessValue <- "2_Bottom_PropertiesTag.ID"
      Appearance <- "2_Bottom_PropertiesTag.ID"
   IOField "valOutputBottom_Category" at 55,25 size 31x26; FormatPattern 99
      ProcessValue <- "2_Bottom_PropertiesTag.Category"
      Appearance <- "2_Bottom_PropertiesTag.ID"
   IOField "valOutputBottom_Message" at 85,25 size 546x26; FormatPattern ??????????????????????????????????????????????????
      ProcessValue <- "2_Bottom_PropertiesTag.Message"
      Appearance <- "2_Bottom_PropertiesTag.ID"
   IOField "valOutputBottom_DateTime" at 630,25 size 201x26
      Appearance <- "2_Bottom_PropertiesTag.ID"
      ProcessValue <- "2_Bottom_PropertiesTag.DateTimeDTL"
   IOField "valOutputBottom_AckDateTime" at 830,25 size 200x26
      Appearance <- "2_Bottom_PropertiesTag.ID"
      ProcessValue <- "2_Bottom_PropertiesTag.AckDateTimeDTL"
*)

(* ===== HMI "HMI_RT_1" =====

ScreenModuleEditorView "fcpEvent_Status_PackMLevent" 745x51
   IOField "valOutputTop_ID" at 0,0 size 56x26; FormatPattern 99999
      ProcessValue <- "1_Top_PropertiesTag.ID"
      Appearance <- "1_Top_PropertiesTag.ID"
   IOField "valOutputTop_Message" at 55,0 size 491x26; FormatPattern ??????????????????????????????????????????????????
      ProcessValue <- "1_Top_PropertiesTag.Message"
      Appearance <- "1_Top_PropertiesTag.ID"
   IOField "valOutputTop_TimeIn" at 545,0 size 200x26
      Appearance <- "1_Top_PropertiesTag.ID"
      ProcessValue <- "1_Top_PropertiesTag.DateTimeDTL"
   IOField "valOutputBottom_ID" at 0,25 size 56x26; FormatPattern 99999
      ProcessValue <- "2_Bottom_PropertiesTag.ID"
      Appearance <- "2_Bottom_PropertiesTag.ID"
   IOField "valOutputBottom_Message" at 55,25 size 491x26; FormatPattern ??????????????????????????????????????????????????
      ProcessValue <- "2_Bottom_PropertiesTag.Message"
      Appearance <- "2_Bottom_PropertiesTag.ID"
   IOField "valOutputBottom_TimeIn" at 545,25 size 200x26
      Appearance <- "2_Bottom_PropertiesTag.ID"
      ProcessValue <- "2_Bottom_PropertiesTag.DateTimeDTL"
*)

(* ===== HMI "HMI_RT_1" =====

ScreenModuleEditorView "fcpOmacStateModel" 1100x550
   GraphicView "pic_btnCmdReset" at 117,396 size 40x40; Picture "Graphic_1"
   GraphicView "pic_btnCmdStart" at 222,179 size 32x32; Picture "media_play_green"
   GraphicView "pic_btnCmdStop" at 330,404 size 27x25; Picture "media_stop_red"
   GraphicView "pic_btnCmdClear" at 633,460 size 40x40; Picture "Graphic_1"
   GraphicView "pic_btnCmdHold" at 650,115 size 32x32; Picture "media_pause"
   TextField "txt_Reset" at 155,400 size 70x32; Text 'Reset'
   TextField "txt_Start" at 203,204 size 70x32; Text 'Start'
   TextField "txt_Stop" at 361,400 size 70x32; Text 'Stop'
   TextField "txt_Clear" at 654,488 size 70x32; Text 'Clear'
   TextField "txt_Hold" at 631,136 size 70x32; Text 'Hold / Start'
   TextField "val_Stopped" at 76,450 size 120x60; Text 'Stopped'
      Appearance <- "i32StateCurrent"
   TextField "val_Resetting" at 76,295 size 120x60; Text 'Resetting'
      Appearance <- "i32StateCurrent"
   TextField "val_Idle" at 76,165 size 120x60; Text 'Idle'
      Appearance <- "i32StateCurrent"
   TextField "val_Starting" at 282,165 size 120x60; Text 'Starting'
      Appearance <- "i32StateCurrent"
   TextField "val_Execute" at 488,165 size 120x60; Text 'Execute'
      Appearance <- "i32StateCurrent"
   TextField "val_Completing" at 694,165 size 120x60; Text 'Completing'
      Appearance <- "i32StateCurrent"
   TextField "val_Complete" at 900,165 size 120x60; Text 'Complete'
      Appearance <- "i32StateCurrent"
   TextField "val_Suspending" at 694,295 size 120x60; Text 'Suspending'
      Appearance <- "i32StateCurrent"
   TextField "val_Suspended" at 488,295 size 120x60; Text 'Suspended'
      Appearance <- "i32StateCurrent"
   TextField "val_Unsuspending" at 282,295 size 120x60; Text 'Un- Suspending'
      Appearance <- "i32StateCurrent"
   TextField "val_Holding" at 694,35 size 120x60; Text 'Holding'
      Appearance <- "i32StateCurrent"
   TextField "val_Held" at 488,35 size 120x60; Text 'Held'
      Appearance <- "i32StateCurrent"
   TextField "val_Unholding" at 282,35 size 120x60; Text 'Un-Holding Un- Holding'
      Appearance <- "i32StateCurrent"
   TextField "val_Aborting" at 900,450 size 120x60; Text 'Aborting'
      Appearance <- "i32StateCurrent"
   TextField "val_Aborted" at 694,450 size 120x60; Text 'Aborted'
      Appearance <- "i32StateCurrent"
   TextField "val_Clearing" at 488,450 size 120x60; Text 'Clearing'
      Appearance <- "i32StateCurrent"
   TextField "val_Stopping" at 282,450 size 120x60; Text 'Stopping'
      Appearance <- "i32StateCurrent"
   TextField "txt_ResettingNotUsed" at 77,295 size 120x60; Text 'Resetting (not used)'
      Visibility <- "i32DisabledStatesInCurrentMode"
   TextField "txt_IdleNotUsed" at 77,165 size 120x60; Text 'Idle (not used)'
      Visibility <- "i32DisabledStatesInCurrentMode"
   TextField "txt_StartingNotUsed" at 283,165 size 120x60; Text 'Starting (not used)'
      Visibility <- "i32DisabledStatesInCurrentMode"
   TextField "txt_CompletingNotUsed" at 695,165 size 120x60; Text 'Completing (not used)'
      Visibility <- "i32DisabledStatesInCurrentMode"
   TextField "txt_CompleteNotUsed" at 901,165 size 120x60; Text 'Complete (not used)'
      Visibility <- "i32DisabledStatesInCurrentMode"
   TextField "txt_SuspendingNotUsed" at 695,295 size 120x60; Text 'Suspending (not used)'
      Visibility <- "i32DisabledStatesInCurrentMode"
   TextField "txt_UnsuspendingNotUsed" at 283,295 size 120x60; Text 'Un-Suspending (not used)'
      Visibility <- "i32DisabledStatesInCurrentMode"
   TextField "txt_HoldingNotUsed" at 695,35 size 120x60; Text 'Holding (not used)'
      Visibility <- "i32DisabledStatesInCurrentMode"
   TextField "txt_HeldNotUsed" at 489,35 size 120x60; Text 'Held (not used)'
      Visibility <- "i32DisabledStatesInCurrentMode"
   TextField "txt_UnholdingNotUsed" at 283,35 size 120x60; Text 'Un-Holding (not used)'
      Visibility <- "i32DisabledStatesInCurrentMode"
   TextField "txt_AbortingNotUsed" at 901,450 size 120x60; Text 'Aborting (not used)'
      Visibility <- "i32DisabledStatesInCurrentMode"
   TextField "txt_ClearingNotUsed" at 489,450 size 120x60; Text 'Clearing (not used)'
      Visibility <- "i32DisabledStatesInCurrentMode"
   TextField "txt_StoppingNotUsed" at 283,450 size 120x60; Text 'Stopping (not used)'
      Visibility <- "i32DisabledStatesInCurrentMode"
   TextField "txt_SuspendedNotUsed" at 489,295 size 120x60; Text 'Suspended (not used) Clearing (not used)'
      Visibility <- "i32DisabledStatesInCurrentMode"

VB script "FaceplateScript_1"
   'Tip:
   ' 1. Use the <CTRL+SPACE> or <CTRL+I> shortcut to open a list of all objects and functions
   ' 2. Write the code using the HMI Runtime object.
   '  Example: HmiRuntime.Screens("Screen_1").
   ' 3. Use the <CTRL+J> shortcut to create an object reference.
   'Write the code as of this position:
*)

(* ===== HMI "HMI_RT_1" =====

HMI tags "Standard-Variablentabelle"
   "bo_FALSE" : Bool, internal

ScreenModuleEditorView "typ_LightStack" 16x58
   Button "val_OutputLightRedStatic" at 0,3 size 16x9; TextOff 'Text'; PictureOff "icn-transparent-15x15px"
      ObjectEnable <- "bo_FALSE"
      Appearance <- "b32_LightStackValue"
   Button "val_OutputLightRedFlashing" at 0,3 size 16x9; TextOff 'Text'; PictureOff "icn-transparent-15x15px"
      Visibility <- "b32_LightStackValue"
      ObjectEnable <- "bo_FALSE"
      Appearance <- "b32_LightStackValue"
   Button "val_OutputLightYellowStatic" at 0,12 size 16x9; TextOff 'Text'; PictureOff "icn-transparent-15x15px"
      ObjectEnable <- "bo_FALSE"
      Appearance <- "b32_LightStackValue"
   Button "val_OutputLightYellowFlashing" at 0,12 size 16x9; TextOff 'Text'; PictureOff "icn-transparent-15x15px"
      Visibility <- "b32_LightStackValue"
      ObjectEnable <- "bo_FALSE"
      Appearance <- "b32_LightStackValue"
   Button "val_OutputLightBlueStatic" at 0,21 size 16x9; TextOff 'Text'; PictureOff "icn-transparent-15x15px"
      ObjectEnable <- "bo_FALSE"
      Appearance <- "b32_LightStackValue"
   Button "val_OutputLightBlueFlashing" at 0,21 size 16x9; TextOff 'Text'; PictureOff "icn-transparent-15x15px"
      Visibility <- "b32_LightStackValue"
      ObjectEnable <- "bo_FALSE"
      Appearance <- "b32_LightStackValue"
   Button "val_OutputLightGreenStatic" at 0,30 size 16x9; TextOff 'Text'; PictureOff "icn-transparent-15x15px"
      ObjectEnable <- "bo_FALSE"
      Appearance <- "b32_LightStackValue"
   Button "val_OutputLightGreenFlashing" at 0,30 size 16x9; TextOff 'Text'; PictureOff "icn-transparent-15x15px"
      Visibility <- "b32_LightStackValue"
      ObjectEnable <- "bo_FALSE"
      Appearance <- "b32_LightStackValue"
   Button "val_OutputLightWhiteStatic" at 0,39 size 16x9; TextOff 'Text'; PictureOff "icn-transparent-15x15px"
      ObjectEnable <- "bo_FALSE"
      Appearance <- "b32_LightStackValue"
   Button "val_OutputLightWhiteFlashing" at 0,39 size 16x9; TextOff 'Text'; PictureOff "icn-transparent-15x15px"
      Visibility <- "b32_LightStackValue"
      ObjectEnable <- "bo_FALSE"
      Appearance <- "b32_LightStackValue"
   Button "fra_LightStackTop" at 0,0 size 16x4; TextOff 'Text'; PictureOff "icn-transparent-15x15px"
   Button "fra_LightStackStand1" at 5,50 size 6x4; TextOff 'Text'; PictureOff "icn-transparent-15x15px"
   Button "fra_LightStackBottom" at 0,47 size 16x4; TextOff 'Text'; PictureOff "icn-transparent-15x15px"
   Button "fra_LightStackStand2" at 0,53 size 16x4; TextOff 'Text'; PictureOff "icn-transparent-15x15px"
*)

(* ===== HMI "HMI_RT_1" =====

ScreenModuleEditorView "fcpOmacStateModel" 1100x550
   GraphicView "pic_btnCmdReset" at 117,396 size 40x40; Picture "Graphic_1"
   GraphicView "pic_btnCmdStart" at 222,179 size 32x32; Picture "media_play_green"
   GraphicView "pic_btnCmdStop" at 330,404 size 27x25; Picture "media_stop_red"
   GraphicView "pic_btnCmdClear" at 633,460 size 40x40; Picture "Graphic_1"
   GraphicView "pic_btnCmdHold" at 650,115 size 32x32; Picture "media_pause"
   TextField "txt_Reset" at 155,400 size 70x32; Text 'Reset'
   TextField "txt_Start" at 203,204 size 70x32; Text 'Start'
   TextField "txt_Stop" at 361,400 size 70x32; Text 'Stop'
   TextField "txt_Clear" at 654,488 size 70x32; Text 'Clear / Reset'
   TextField "txt_Hold" at 631,136 size 70x32; Text 'Hold / Start'
   TextField "val_Stopped" at 76,450 size 120x60; Text 'Stopped'
      Appearance <- "i32StateCurrent"
   TextField "val_Resetting" at 76,295 size 120x60; Text 'Resetting'
      Appearance <- "i32StateCurrent"
   TextField "val_Idle" at 76,165 size 120x60; Text 'Idle'
      Appearance <- "i32StateCurrent"
   TextField "val_Starting" at 282,165 size 120x60; Text 'Starting'
      Appearance <- "i32StateCurrent"
   TextField "val_Execute" at 488,165 size 120x60; Text 'Execute'
      Appearance <- "i32StateCurrent"
   TextField "val_Completing" at 694,165 size 120x60; Text 'Completing'
      Appearance <- "i32StateCurrent"
   TextField "val_Complete" at 900,165 size 120x60; Text 'Complete'
      Appearance <- "i32StateCurrent"
   TextField "val_Suspending" at 694,295 size 120x60; Text 'Suspending'
      Appearance <- "i32StateCurrent"
   TextField "val_Suspended" at 488,295 size 120x60; Text 'Suspended'
      Appearance <- "i32StateCurrent"
   TextField "val_Unsuspending" at 282,295 size 120x60; Text 'Un- Suspending'
      Appearance <- "i32StateCurrent"
   TextField "val_Holding" at 694,35 size 120x60; Text 'Holding'
      Appearance <- "i32StateCurrent"
   TextField "val_Held" at 488,35 size 120x60; Text 'Held'
      Appearance <- "i32StateCurrent"
   TextField "val_Unholding" at 282,35 size 120x60; Text 'Un-Holding Un- Holding'
      Appearance <- "i32StateCurrent"
   TextField "val_Aborting" at 900,450 size 120x60; Text 'Aborting'
      Appearance <- "i32StateCurrent"
   TextField "val_Aborted" at 694,450 size 120x60; Text 'Aborted'
      Appearance <- "i32StateCurrent"
   TextField "val_Clearing" at 488,450 size 120x60; Text 'Clearing'
      Appearance <- "i32StateCurrent"
   TextField "val_Stopping" at 282,450 size 120x60; Text 'Stopping'
      Appearance <- "i32StateCurrent"
   TextField "txt_ResettingNotUsed" at 77,295 size 120x60; Text 'Resetting (not used)'
      Visibility <- "i32DisabledStatesInCurrentMode"
   TextField "txt_IdleNotUsed" at 77,165 size 120x60; Text 'Idle (not used)'
      Visibility <- "i32DisabledStatesInCurrentMode"
   TextField "txt_StartingNotUsed" at 283,165 size 120x60; Text 'Starting (not used)'
      Visibility <- "i32DisabledStatesInCurrentMode"
   TextField "txt_CompletingNotUsed" at 695,165 size 120x60; Text 'Completing (not used)'
      Visibility <- "i32DisabledStatesInCurrentMode"
   TextField "txt_CompleteNotUsed" at 901,165 size 120x60; Text 'Complete (not used)'
      Visibility <- "i32DisabledStatesInCurrentMode"
   TextField "txt_SuspendingNotUsed" at 695,295 size 120x60; Text 'Suspending (not used)'
      Visibility <- "i32DisabledStatesInCurrentMode"
   TextField "txt_UnsuspendingNotUsed" at 283,295 size 120x60; Text 'Un-Suspending (not used)'
      Visibility <- "i32DisabledStatesInCurrentMode"
   TextField "txt_HoldingNotUsed" at 695,35 size 120x60; Text 'Holding (not used)'
      Visibility <- "i32DisabledStatesInCurrentMode"
   TextField "txt_HeldNotUsed" at 489,35 size 120x60; Text 'Held (not used)'
      Visibility <- "i32DisabledStatesInCurrentMode"
   TextField "txt_UnholdingNotUsed" at 283,35 size 120x60; Text 'Un-Holding (not used)'
      Visibility <- "i32DisabledStatesInCurrentMode"
   TextField "txt_AbortingNotUsed" at 901,450 size 120x60; Text 'Aborting (not used)'
      Visibility <- "i32DisabledStatesInCurrentMode"
   TextField "txt_ClearingNotUsed" at 489,450 size 120x60; Text 'Clearing (not used)'
      Visibility <- "i32DisabledStatesInCurrentMode"
   TextField "txt_StoppingNotUsed" at 283,450 size 120x60; Text 'Stopping (not used)'
      Visibility <- "i32DisabledStatesInCurrentMode"
   TextField "txt_SuspendedNotUsed" at 489,295 size 120x60; Text 'Suspended (not used) Clearing (not used)'
      Visibility <- "i32DisabledStatesInCurrentMode"

VB script "FaceplateScript_1"
   'Tip:
   ' 1. Use the <CTRL+SPACE> or <CTRL+I> shortcut to open a list of all objects and functions
   ' 2. Write the code using the HMI Runtime object.
   '  Example: HmiRuntime.Screens("Screen_1").
   ' 3. Use the <CTRL+J> shortcut to create an object reference.
   'Write the code as of this position:
*)

(* ===== HMI "HMI_RT_1" =====

ScreenModuleEditorView "ParetoFacePlate" 1200x200
   IOField "Field_alarmID" at 126,76 size 55x32; FormatPattern 9999
      ProcessValue <- "Property_1.alarmID"
   IOField "Field_alarmMessage" at 191,76 size 334x32; FormatPattern ????????????????????????????????????????
      ProcessValue <- "Property_1.alarmMessage"
   IOField "Field_TimesOccurred" at 536,76 size 41x32; FormatPattern 99
      ProcessValue <- "Property_1.timesOccurred"
   IOField "Field_totalDowntime" at 587,76 size 59x32; FormatPattern 999.99
      ProcessValue <- "Property_1.totalDowntime"
   IOField "Field_MTTR" at 657,76 size 59x32; FormatPattern 999.99
      ProcessValue <- "Property_1.MTTR"
   IOField "Field_PercentageOccurred" at 727,76 size 47x32; FormatPattern 99.9
      ProcessValue <- "Property_1.percentageOccurred"
*)

(* ===== HMI "HMI_RT_1" =====
system functions are stored by id; their names below are inferred from use
connection "HMI_TP1200_Connection": ETHERNET, S7_1500_OMS
